// TIA Portal project "CHM_BORDEIRA_20190721" (V15)
// Frazer-Nash Consultancy Edits

(* hardware
DEVICE "SCALANCE X005"  SCALANCE X-Station
   slot 0: "SCALANCE X rack"  Rail
   slot 0: "Switch_1"  6GK5 008-0BA00-1AB2  V1.0
DEVICE "RIO 2/RIOCP-2T-ET 200iSP"  ET 200iSP station
   slot 0: "RIO 2 / RIOCP-2T"  Rail
   slot 2: "RIO 2 / RIOCP-2T - 5KF1 - IF Module"  ET200iSP  6ES7 152-1AA00-0AB0  V2.0
   slot 4: "6KF1 - 8DI x NAMUR"  8DI x NAMUR  6ES7 131-7RF00-0AB0
   slot 5: "7KF1 - 8DI x NAMUR"  8DI x NAMUR  6ES7 131-7RF00-0AB0
   slot 6: "8KF1 - 8DI x NAMUR"  8DI x NAMUR  6ES7 131-7RF00-0AB0
   slot 7: "9KF1 - 4DO x 23.1VDC / 20mA SD 'H'"  4DO x 23.1VDC / 20mA SD 'H'  6ES7 132-7RD01-0AB0
   slot 8: "10KF1 - 4AI x 2WIRE HART"  4AI x 2WIRE HART  6ES7 134-7TD00-0AB0
   slot 9: "11KF1 - 4AI x 2WIRE HART"  4AI x 2WIRE HART  6ES7 134-7TD00-0AB0
   slot 10: "12KF1 - 4AI x 2WIRE HART"  4AI x 2WIRE HART  6ES7 134-7TD00-0AB0
   slot 11: "13KF1 - 4AI x 2WIRE HART"  4AI x 2WIRE HART  6ES7 134-7TD00-0AB0
DEVICE "ET 200SP station_1"  ET 200SP-Station
   slot 0: "Rack_1"  Rack  6ES5 710-8MAx1
   slot 1: "Rack 1 - IGG PLC - 15KF2"  CPU 1510SP-1 PN  6ES7 510-1DJ01-0AB0  V2.1
   slot 2: "16KF1 - DI 16x24VDC ST_1"  DI 16x24VDC ST  6ES7 131-6BH00-0BA0  V1.1
      slot 1: "16KF1 - DI 16x24VDC ST_1"  DI 16x24VDC ST
   slot 3: "18KF1 - DI 16x24VDC ST_2"  DI 16x24VDC ST  6ES7 131-6BH00-0BA0  V1.1
      slot 1: "18KF1 - DI 16x24VDC ST_2"  DI 16x24VDC ST
   slot 4: "23KF1 - DQ 16x24VDC/0.5A ST_1"  DQ 16x24VDC/0.5A ST  6ES7 132-6BH00-0BA0  V1.1
      slot 1: "23KF1 - DQ 16x24VDC/0.5A ST_1"  DQ 16x24VDC/0.5A ST
   slot 5: "29KF1 - AI 8xI 2-,4-wire BA_1"  AI 8xI 2-,4-wire BA  6ES7 134-6GF00-0AA1  V1.0
      slot 1: "29KF1 - AI 8xI 2-,4-wire BA_1"  AI 8xI 2-,4-wire BA
   slot 6: "31KF1 - AI 8xI 2-,4-wire BA_2"  AI 8xI 2-,4-wire BA  6ES7 134-6GF00-0AA1  V1.0
      slot 1: "31KF1 - AI 8xI 2-,4-wire BA_2"  AI 8xI 2-,4-wire BA
   slot 7: "35KF1 - AQ 4xU/I ST_1"  AQ 4xU/I ST  6ES7 135-6HD00-0BA1  V1.1
      slot 1: "35KF1 - AQ 4xU/I ST_1"  AQ 4xU/I ST
   slot 8: "Server module_1"  Server module  6ES7 193-6PA00-0AA0  V1.0
      slot 1: "Server module_1"  Server module
   slot 127: "PROFINET BusAdapter CU"  BA 2xRJ45  6ES7 193-6AR00-0AA0  V0.0
      slot 32769: "Port_1"  6ES7 193-6AR00-0AA0
      slot 32770: "Port_2"  6ES7 193-6AR00-0AA0
DEVICE "ET 200SP station_2"  ET 200SP-Station
   slot 0: "Rack_2"  Rack  6ES5 710-8MAx1
   slot 1: "Rack 2 - BC PLC - 15KF3"  CPU 1510SP-1 PN  6ES7 510-1DJ01-0AB0  V2.1
   slot 2: "19KF1 - DI 16x24VDC ST_1"  DI 16x24VDC ST  6ES7 131-6BH00-0BA0  V1.1
      slot 1: "19KF1 - DI 16x24VDC ST_1"  DI 16x24VDC ST
   slot 3: "21KF1 - DI 16x24VDC ST_2"  DI 16x24VDC ST  6ES7 131-6BH00-0BA0  V1.1
      slot 1: "21KF1 - DI 16x24VDC ST_2"  DI 16x24VDC ST
   slot 4: "25KF1 - DQ 16x24VDC/0.5A ST_1"  DQ 16x24VDC/0.5A ST  6ES7 132-6BH00-0BA0  V1.1
      slot 1: "25KF1 - DQ 16x24VDC/0.5A ST_1"  DQ 16x24VDC/0.5A ST
   slot 5: "33KF1 - AI 8xI 2-,4-wire BA_1"  AI 8xI 2-,4-wire BA  6ES7 134-6GF00-0AA1  V1.0
      slot 1: "33KF1 - AI 8xI 2-,4-wire BA_1"  AI 8xI 2-,4-wire BA
   slot 6: "37KF1 - AQ 4xU/I ST_1"  AQ 4xU/I ST  6ES7 135-6HD00-0BA1  V1.1
      slot 1: "37KF1 - AQ 4xU/I ST_1"  AQ 4xU/I ST
   slot 7: "Server module_1"  Server module  6ES7 193-6PA00-0AA0  V1.0
      slot 1: "Server module_1"  Server module
   slot 127: "PROFINET BusAdapter CU"  BA 2xRJ45  6ES7 193-6AR00-0AA0  V0.0
      slot 32769: "Port_1"  6ES7 193-6AR00-0AA0
      slot 32770: "Port_2"  6ES7 193-6AR00-0AA0
DEVICE "S71500/ET200MP station_1"  S7-1500 station
   slot 0: "Rail_0"  Rack  6ES7 590-1***0-0AA0
   slot 1: "Rack 3 - GCU & BWT PLC - 7KF2"  CPU 1516F-3 PN/DP  6ES7 516-3FN01-0AB0  V2.1
      slot 3: "CPU display_1"  6ES7591-1BA00-0AA0
   slot 2: "8KF1 - DI 32x24VDC HF_1"  DI 32x24VDC HF  6ES7 521-1BL00-0AB0  V2.1
   slot 3: "12KF1 - DQ 32x24VDC/0.5A HF_1"  DQ 32x24VDC/0.5A HF  6ES7 522-1BL01-0AB0  V1.0
   slot 4: "16KF1 - AI 8xU/I HF_2"  AI 8xU/I HF  6ES7 531-7NF00-0AB0  V1.0
   slot 5: "18KF1 - AI 8xU/I HF_1"  AI 8xU/I HF  6ES7 531-7NF00-0AB0  V1.0
   slot 6: "20KF1 - AQ 4xU/I HF_1"  AQ 4xU/I HF  6ES7 532-5ND00-0AB0  V1.0
DEVICE "RIO 1/RIOCP-3T-ET 200iSP"  ET 200iSP station
   slot 0: "RIO 1 / RIOCP-3T"  Rail
   slot 2: "RIO 1 / RIOCP-3T - 5KF1 - IF Module"  ET200iSP  6ES7 152-1AA00-0AB0  V2.0
   slot 4: "6KF1 - 8DI x NAMUR_1"  8DI x NAMUR  6ES7 131-7RF00-0AB0
   slot 5: "7KF1 - 8DI x NAMUR_2"  8DI x NAMUR  6ES7 131-7RF00-0AB0
   slot 6: "8KF1 - 8DI x NAMUR_3"  8DI x NAMUR  6ES7 131-7RF00-0AB0
   slot 7: "9KF1 - 8DI x NAMUR_4"  8DI x NAMUR  6ES7 131-7RF00-0AB0
   slot 8: "10KF1 - 4DO x 23.1VDC / 20mA SD 'H'_1"  4DO x 23.1VDC / 20mA SD 'H'  6ES7 132-7RD01-0AB0
   slot 9: "11KF1 - 4DO x 23.1VDC / 20mA SD 'H'_2"  4DO x 23.1VDC / 20mA SD 'H'  6ES7 132-7RD01-0AB0
   slot 10: "12KF1 - 4AI x 2WIRE HART_1"  4AI x 2WIRE HART  6ES7 134-7TD00-0AB0
   slot 11: "13KF1 - 4AI x 2WIRE HART_2"  4AI x 2WIRE HART  6ES7 134-7TD00-0AB0
   slot 12: "14KF1 - 4AI x 2WIRE HART_1"  4AI x 2WIRE HART  6ES7 134-7TD00-0AB0
   slot 13: "15KF1 - 4AI x 2WIRE HART_2"  4AI x 2WIRE HART  6ES7 134-7TD00-0AB0
   slot 14: "16KF1 - 4AI x 2WIRE HART_3"  4AI x 2WIRE HART  6ES7 134-7TD00-0AB0
   slot 15: "17KF1 - 4AI x 2WIRE HART_4"  4AI x 2WIRE HART  6ES7 134-7TD00-0AB0
   slot 16: "Standby modules_1"  Standby modules  6ES7 138-7AA00-0AA0
DEVICE "RIO 3/RIOCP-2T-ET 200iSP"  ET 200iSP station
   slot 0: "RIO 3 / RIOCP-2T"  Rail
   slot 2: "RIO 3 / RIOCP-2T - 5KF1 - IF Module"  ET200iSP  6ES7 152-1AA00-0AB0  V2.0
   slot 4: "6KF1 - 8DI x NAMUR"  8DI x NAMUR  6ES7 131-7RF00-0AB0
   slot 5: "7KF1 - 8DI x NAMUR"  8DI x NAMUR  6ES7 131-7RF00-0AB0
   slot 6: "8KF1 - 8DI x NAMUR"  8DI x NAMUR  6ES7 131-7RF00-0AB0
   slot 7: "9KF1 - 4DO x 23.1VDC / 20mA SD 'H'"  4DO x 23.1VDC / 20mA SD 'H'  6ES7 132-7RD01-0AB0
   slot 8: "10KF1 - 4AI x 2WIRE HART_1"  4AI x 2WIRE HART  6ES7 134-7TD00-0AB0
   slot 9: "11KF1 - 4AI x 2WIRE HART"  4AI x 2WIRE HART  6ES7 134-7TD00-0AB0
   slot 10: "12KF1 - 4AI x 2WIRE HART"  4AI x 2WIRE HART  6ES7 134-7TD00-0AB0
   slot 11: "13KF1 - 4AI x 2WIRE HART"  4AI x 2WIRE HART  6ES7 134-7TD00-0AB0
DEVICE "RIO 4/RIOCP-2T-ET 200iSP"  ET 200iSP station
   slot 0: "RIO 4 / RIOCP-2T"  Rail
   slot 2: "RIO 4 / RIOCP-2T - 5KF1 - IF Module"  ET200iSP  6ES7 152-1AA00-0AB0  V2.0
   slot 4: "6KF1 - 8DI x NAMUR"  8DI x NAMUR  6ES7 131-7RF00-0AB0
   slot 5: "7KF1 - 8DI x NAMUR"  8DI x NAMUR  6ES7 131-7RF00-0AB0
   slot 6: "8KF1 - 8DI x NAMUR"  8DI x NAMUR  6ES7 131-7RF00-0AB0
   slot 7: "9KF1 - 4DO x 23.1VDC / 20mA SD 'H'"  4DO x 23.1VDC / 20mA SD 'H'  6ES7 132-7RD01-0AB0
   slot 8: "10KF1 - 4AI x 2WIRE HART_1"  4AI x 2WIRE HART  6ES7 134-7TD00-0AB0
   slot 9: "11KF1 - 4AI x 2WIRE HART_1"  4AI x 2WIRE HART  6ES7 134-7TD00-0AB0
   slot 10: "12KF1 - 4AI x 2WIRE HART"  4AI x 2WIRE HART  6ES7 134-7TD00-0AB0
   slot 11: "13KF1 - 4AI x 2WIRE HART"  4AI x 2WIRE HART  6ES7 134-7TD00-0AB0
DEVICE "RIO 5/RIOCP-2T-ET 200iSP"  ET 200iSP station
   slot 0: "RIO 5 / RIOCP-2T"  Rail
   slot 2: "RIO 5 / RIOCP-2T - 5KF1 - IF Module"  ET200iSP  6ES7 152-1AA00-0AB0  V2.0
   slot 4: "6KF1 - 8DI x NAMUR_1"  8DI x NAMUR  6ES7 131-7RF00-0AB0
   slot 5: "7KF1 - 8DI x NAMUR_2"  8DI x NAMUR  6ES7 131-7RF00-0AB0
   slot 6: "8KF1 - 8DI x NAMUR_3"  8DI x NAMUR  6ES7 131-7RF00-0AB0
   slot 7: "9KF1 - 4DO x 23.1VDC / 20mA SD 'H'_1"  4DO x 23.1VDC / 20mA SD 'H'  6ES7 132-7RD01-0AB0
   slot 8: "10KF1 - 4AI x 2WIRE HART_1"  4AI x 2WIRE HART  6ES7 134-7TD00-0AB0
   slot 9: "11KF1- 4AI x 2WIRE HART_1"  4AI x 2WIRE HART  6ES7 134-7TD00-0AB0
   slot 10: "12KF1 - 4AI x 2WIRE HART_2"  4AI x 2WIRE HART  6ES7 134-7TD00-0AB0
   slot 11: "13KF1 - 4AI x 2WIRE HART_3"  4AI x 2WIRE HART  6ES7 134-7TD00-0AB0
DEVICE "RIO 7/RIOCP-1T-ET 200iSP"  ET 200iSP station
   slot 0: "RIO 7/ RIOCP-1T"  Rail
   slot 2: "RIO 7 / RIOCP-1T - 5KF1 - IF Module"  ET200iSP  6ES7 152-1AA00-0AB0  V2.0
   slot 4: "6KF1 - 8DI x NAMUR"  8DI x NAMUR  6ES7 131-7RF00-0AB0
   slot 5: "7KF1 - 8DI x NAMUR"  8DI x NAMUR  6ES7 131-7RF00-0AB0
   slot 6: "8KF1 - 4DO x 23.1VDC / 20mA SD 'H'_1"  4DO x 23.1VDC / 20mA SD 'H'  6ES7 132-7RD01-0AB0
   slot 7: "9KF1 - 4AI x 2WIRE HART_1"  4AI x 2WIRE HART  6ES7 134-7TD00-0AB0
   slot 8: "10KF1 - 4AI x 2WIRE HART"  4AI x 2WIRE HART  6ES7 134-7TD00-0AB0
   slot 9: "11KF1 - 4AI x 2WIRE HART"  4AI x 2WIRE HART  6ES7 134-7TD00-0AB0
DEVICE "RIO 6/RIOCP-2T-ET 200iSP"  ET 200iSP station
   slot 0: "RIO 6 / RIOCP-2T"  Rail
   slot 2: "RIO 6 / RIOCP-2T - 5KF1 - IF Module"  ET200iSP  6ES7 152-1AA00-0AB0  V2.0
   slot 4: "6KF1 - 8DI x NAMUR_1"  8DI x NAMUR  6ES7 131-7RF00-0AB0
   slot 5: "7KF1 - 8DI x NAMUR_2"  8DI x NAMUR  6ES7 131-7RF00-0AB0
   slot 6: "8KF1 - 8DI x NAMUR_3"  8DI x NAMUR  6ES7 131-7RF00-0AB0
   slot 7: "9KF1 - 4DO x 23.1VDC / 20mA SD 'H'_1"  4DO x 23.1VDC / 20mA SD 'H'  6ES7 132-7RD01-0AB0
   slot 8: "10KF1 - 4AI x 2WIRE HART_1"  4AI x 2WIRE HART  6ES7 134-7TD00-0AB0
   slot 9: "11KF1- 4AI x 2WIRE HART_1"  4AI x 2WIRE HART  6ES7 134-7TD00-0AB0
   slot 10: "12KF1 - 4AI x 2WIRE HART_2"  4AI x 2WIRE HART  6ES7 134-7TD00-0AB0
   slot 11: "13KF1 - 4AI x 2WIRE HART_3"  4AI x 2WIRE HART  6ES7 134-7TD00-0AB0
DEVICE "IGG HMI"  TP1500 Comfort
   slot 0: "IGG HMI"  TP1500 Comfort  6AV2 124-0QC02-0AX0  15.0.0.0
   slot 1: "HMI_RT_1"  TP1500 Comfort  6AV2 124-0QC02-0AX0  15.0.0.0
   slot 5: "IGG HMI.IE_CP_1"  PROFINET Interface  15.0.0.0
      slot 1: "PROFINET Interface_1"  PROFINET Interface
         slot 1: "Port_1"  Port
         slot 2: "Port_2"  Port
   slot 6: "IGG HMI.IE_CP_2"  PROFINET Interface  15.0.0.0
      slot 1: "PROFINET Interface_GBit"  PROFINET Interface
         slot 1: "Port_1"  Port
   slot 7: "IGG HMI.MPI/DP_CP_1"  MPI/DP Interface  15.0.0.0
DEVICE "CCR HMI"  TP1200 Comfort
   slot 0: "CCR HMI"  TP1200 Comfort  6AV2 124-0MC01-0AX0  15.0.0.0
   slot 1: "HMI_RT_4"  TP1200 Comfort  6AV2 124-0MC01-0AX0  15.0.0.0
   slot 5: "CCR HMI._CP_1"  PROFINET Interface  15.0.0.0
      slot 1: "PROFINET Interface_1"  PROFINET Interface
         slot 1: "Port_1"  Port
         slot 2: "Port_2"  Port
   slot 7: "CCR HMI.I/DP_CP_1"  MPI/DP Interface  15.0.0.0
DEVICE "Bridge HMI"  KTP400 Comfort
   slot 0: "Bridge HMI"  KTP400 Comfort  6AV2 124-2DC01-0AX0  15.0.0.0
   slot 1: "HMI_RT_2"  KTP400 Comfort  6AV2 124-2DC01-0AX0  15.0.0.0
   slot 5: "Bridge HMI.1"  PROFINET Interface  15.0.0.0
      slot 1: "PROFINET Interface_1"  PROFINET Interface
         slot 1: "Port_1"  Port
   slot 7: "Bridge HMI._CP_1"  MPI/DP Interface  15.0.0.0
DEVICE "GSD device_1"  GSD.Device.PN
   slot 0: "Rack"  Rack  V1.0
   slot 0: "WBT"  Serial  HD674-A006
      slot 0: "Submodule V1"  Submodule V1
      slot 1: "I"  I
         slot 1: "P1"  P1
         slot 2: "P2"  P2
   slot 1: "IO"  Module  12345-0040-M
      slot 0: "Module"  Module
*)

// ===== PLC "Rack 1 - IGG PLC - 15KF2"  CPU 1510SP-1 PN =====

VAR_GLOBAL   // PLC tag table "Default tag table"
   "System_Byte" AT %MB1 : Byte;
   "FirstScan" AT %M1.0 : Bool;
   "DiagStatusUpdate" AT %M1.1 : Bool;
   "AlwaysTRUE" AT %M1.2 : Bool;
   "AlwaysFALSE" AT %M1.3 : Bool;
   "Clock_Byte" AT %MB0 : Byte;
   "Clock_10Hz" AT %M0.0 : Bool;
   "Clock_5Hz" AT %M0.1 : Bool;
   "Clock_2.5Hz" AT %M0.2 : Bool;
   "Clock_2Hz" AT %M0.3 : Bool;
   "Clock_1.25Hz" AT %M0.4 : Bool;
   "Clock_1Hz" AT %M0.5 : Bool;
   "Clock_0.625Hz" AT %M0.6 : Bool;
   "Clock_0.5Hz" AT %M0.7 : Bool;
   "IGG E-Stop Healthy" AT %I0.0 : Bool;   // S2-8K1
   "CA Blower Ready" AT %I0.1 : Bool;   // E139-MCCP/6TA1
   "Fuel Pump 1 Tripped" AT %I0.2 : Bool;   // E500A-MCCP/7Q2
   "Fuel Pump 2 Tripped" AT %I0.3 : Bool;   // E500B-MCCP/7Q3
   "Fuel Pump 1 Enabled" AT %I0.4 : Bool;   // E500A-MCCP/9Q1
   "Fuel Pump 2 Enabled" AT %I0.5 : Bool;   // E500B-MCCP/9Q2
   "IG Supply Valve Opened" AT %I0.6 : Bool;   // CV401-16B1
   "IG Supply Valve Closed" AT %I0.7 : Bool;   // CV401-16B1
   "DTB Valve Opened" AT %I1.0 : Bool;   // CV321-17B1
   "DTB Valve Closed" AT %I1.1 : Bool;   // CV321-17B1
   "CSW Drain Valve Opened" AT %I1.2 : Bool;   // CV322-17B2
   "CSW Drain Valve Closed" AT %I1.3 : Bool;   // CV322-17B2
   "CSW Valve Open" AT %I1.4 : Bool;   // CV311-17B3
   "CSW Valve Closed" AT %I1.5 : Bool;   // CV311-17B3
   "Flue Gas Scrubber CSW Valve Opened" AT %I1.6 : Bool;   // CV312-17B4
   "Flue Gas Scrubber CSW Valve Closed" AT %I1.7 : Bool;   // CV312-17B4
   "BC PLC Power Healthy" AT %I2.0 : Bool;   // -15Q4
   "IGG Vent Power Healthy" AT %I2.1 : Bool;   // -6Q2
   "MCC Vent Power Healthy" AT %I2.2 : Bool;   // -MCCP/8Q4
   "7T1 Power Healthy" AT %I2.3 : Bool;   // -7T1 Controls Power
   "7T2 Power Healthy" AT %I2.4 : Bool;   // -7T2 IGG Power
   "7T3 Power Healthy" AT %I2.5 : Bool;   // -7T3 BC Power
   "Maintained 24V Power" AT %I2.6 : Bool;   // -7Q4
   "Safety System Interlock" AT %I2.7 : Bool;   // Safety interlock
   "Cargo Blanketing IG Supply Valve Open" AT %I3.0 : Bool;   // CV431-25QM8
   "Cargo Blanketing IG Supply Valve Close" AT %I3.1 : Bool;   // CV431-25QM8
   "BWTS IG Supply Valve Open" AT %I3.2 : Bool;   // CV432-25QM8
   "BWTS IG Supply Valve Close" AT %I3.3 : Bool;   // CV432-25QM8
   "CA Blower Running" AT %I3.4 : Bool;   // E139-MCCP/6TA1
   "VSD Fault" AT %I3.5 : Bool;   // E139-MCCP/6TA1
   "Correct Phase Rotation" AT %I3.6 : Bool;   // -MCCP/5PG1
   "R1_SPR_DI_3_7" AT %I3.7 : Bool;   // Spare input
   "CA Pressure PIT102" AT %IW112 : Int;   // PIT102-29B1
   "IG Temp" AT %IW114 : Int;   // TIT401-29B2
   "IG Outlet Pressure PIT402" AT %IW116 : Int;   // PIT402-29B3
   "IG Vent Valve Position Feedback" AT %IW118 : Int;   // CV403-29B4
   "CA Blower RPM" AT %IW120 : Int;   // E139-6TA1
   "CA Blower Current" AT %IW122 : Int;   // E139-6TA1
   "FW Bulk Tank Level Transmitter" AT %IW124 : Int;   // LIT305
   "Atm Oxygen Content 1" AT %IW128 : Int;   // Crowcon Atmospheric Sensors-31B1
   "Atm Oxygen Content 2" AT %IW130 : Int;   // Crowcon Atmospheric Sensors-31B2
   "R1_SPR_AI_132" AT %IW132 : Int;   // Spare
   "Shell CSW Temp TIT315" AT %IW134 : Int;   // TIT315-31B4
   "Inlet CSW Temp TIT319" AT %IW136 : Int;   // TIT319-32B1
   "Outlet CSW Temp TIT360" AT %IW138 : Int;   // TIT360-32B2
   "Inlet CSW Pressure PIT359" AT %IW140 : Int;   // PIT359-32B3
   "Outlet CSW Pressure PIT316" AT %IW142 : Int;   // PIT316-32B4
   "Fuel Pump 1 Control" AT %Q0.0 : Bool;   // E500-MCCP/9Q1
   "Fuel Pump 2 Control" AT %Q0.1 : Bool;   // E500-MCCP/9Q1
   "CA Blower Control" AT %Q0.2 : Bool;   // E139-MCCP/6TA1
   "CSW Inlet Valves Control" AT %Q0.3 : Bool;   // CV311/CV312-23QM1
   "CSW Drain Valves Control" AT %Q0.4 : Bool;   // CV321/CV322-23QM2
   "IG Supply Valve Control" AT %Q0.5 : Bool;   // CV401
   "R1_SPR_DQ_1_0" AT %Q1.0 : Bool;   // Spare input
   "Atmospheric Alarm" AT %Q1.1 : Bool;   // -24K2
   "IGG Shutdown Alarm Active" AT %Q1.2 : Bool;   // -24K3
   "IGG Warning Alarm Active" AT %Q1.3 : Bool;   // -24K4
   "IGG Running" AT %Q1.4 : Bool;   // -24PF1
   "Shutdown Alarm" AT %Q1.5 : Bool;   // -24PF2
   "Warning Alarm" AT %Q1.6 : Bool;   // -24PF3
   "Buzzer" AT %Q1.7 : Bool;   // -24PF4
   "Vent Valve Position Control" AT %QW98 : Int;   // CV403-35QN1
   "R1_SPR_AI_126" AT %IW126 : Int;   // Spare input
   "Cargo Blanketing/BWTS Valve Control" AT %Q0.6 : Bool;   // CV431/432-25QM8
   "R1_SPR_DQ_0_7" AT %Q0.7 : Bool;   // Spare input
   "CA Blower Speed Control" AT %QW100 : Word;   // E139-MCCP/6TA1
   "R1_SPR_AQ_102" AT %QW102 : Word;   // Spare output
   "R1_SPR_AQ_104" AT %QW104 : Word;   // Spare output
   "db_time_sync_time_system_READ" AT %M2.0 : LDT;
   "db_time_sync_time_local_READ" AT %M4.0 : LDT;
   "TimeRetVal1" AT %MW8 : Int;
   "RESET_STEP" AT %M12.0 : Bool;
   "IGG_ALARM_ACKNLG_1" AT %MW12 : Word;   // %MW12.DBX0.0
   "IGG_ALARM_ACKNLG_2" AT %MW14 : Word;
   "IGG_ALARM_ACKNLG_3" AT %MW16 : Word;
   "IGG_ALARM_ACKNLG_4" AT %MW18 : Word;
   "IGG_ALARM_ACKNLG_5" AT %MW20 : Word;
   "IGG_ALARM_ACKNLG_6" AT %MW22 : Word;
   "BC_ALARM_ACKNLG_1" AT %MW24 : Word;
   "BC_ALARM_ACKNLG_2" AT %MW26 : Word;
   "BC_ALARM_ACKNLG_3" AT %MW28 : Word;
   "BC_ALARM_ACKNLG_4" AT %MW30 : Word;
   "BC_ALARM_ACKNLG_5" AT %MW32 : Word;
   "BC_ALARM_ACKNLG_6" AT %MW34 : Word;
   "Tag_1" AT %M233.3 : Bool;
   "Tag_2" AT %M233.4 : Bool;
   "Tag_3" AT %M233.5 : Bool;
   "Tag_4" AT %M233.6 : Bool;
   "Tag_5" AT %M233.7 : Bool;
END_VAR

TYPE "AI_Data"
VERSION : 0.1
   STRUCT
      RAW_MIN : Int;   // Raw minimum value from AI card
      RAW_MAX : Int := 27648;   // Raw maximum value from AI card
      NORM : Real;   // Normalised real value
      ENG_MIN : Real;   // Engineering units minimum value
      ENG_MAX : Real := 100.0;   // Engineering units maximum value
   END_STRUCT;
END_TYPE

TYPE "AQ_Data"
VERSION : 0.1
   STRUCT
      ENG_MIN : Real;   // Engineering units minimum value
      ENG_MAX : Real := 100.0;   // Engineering units maximum value
      NORM : Real;   // Normalised real value
      RAW_MIN : Int;   // Raw minimum value from AQ card
      RAW_MAX : Int := 27648;   // Raw maximum value from AQ card
   END_STRUCT;
END_TYPE

// folder: 10 - 19 IO & Processing

DATA_BLOCK "Alarm beacon handling_DB"   // DB1
{ S7_Optimized_Access := 'TRUE' }
VERSION : 0.1
// stored: InstanceOfName Alarm beacon handling
"Alarm beacon handling"
BEGIN
END_DATA_BLOCK

DATA_BLOCK "Date_And_Time_Data"   // DB3
{ S7_Optimized_Access := 'TRUE' }
VERSION : 0.1
   VAR
      SYSTEM_TIME : DTL;
      LOCAL_TIME : DTL;
      HMI_INPUT_FIELD_TIME_IGG : DTL;
      SYNCH_HMI_CLOCK_IGG : Bool;
      GET_TIME_IGG : Bool;
      HMI_INPUT_FIELD_TIME_CCR : DTL;
      SYNCH_HMI_CLOCK_CCR : Bool;
      GET_TIME_CCR : Bool;
   END_VAR
BEGIN
END_DATA_BLOCK

DATA_BLOCK "10_DI_Data"   // DB10
TITLE = Digital Input Data
{ S7_Optimized_Access := 'TRUE' }
AUTHOR : JRS
VERSION : 0.1
// Processed data for code use
   VAR
      IGG_ESTOP_OK : Bool;   // IGG E-Stop healthy (S2-8K1)
      BC_PLC_PWR_OK : Bool;   // BC PLC Power healthy
      IGG_VNT_PWR_OK : Bool;   // IGG Vent power healthy
      MCC_VNT_PWR_OK : Bool;   // MCC Vent power healthy
      "7T1_PWR_OK" : Bool;   // 7T1 Power healthy
      "7T2_PWR_OK" : Bool;   // 7T2 Power healthy
      "7T3_PWR_OK" : Bool;   // 7T3 Power healthy
      MAINTD_24VDC_PWR_OK : Bool;   // Maintained 24V power
      SFTY_SYS_IL : Bool;   // Safety system interlock
      R1_SPR_DI_3_7 : Bool;   // Spare input
      MCCP_5PG1_OK : Bool;   // Correct phase rotation
      CV311_OPN : Bool;   // CSW Valve Open
      CV311_CLSD : Bool;   // CSW Valve Closed
      CV312_OPN : Bool;   // Flue Gas Scrubber CSW valve open
      CV312_CLSD : Bool;   // Flue gas scrubber CSW valve closed
      CV321_OPN : Bool;   // DTB valve open
      CV321_CLSD : Bool;   // DTB valve closed
      CV322_OPN : Bool;   // CSW Drain valve open
      CV322_CLSD : Bool;   // CSW drain valve closed
      CV401_OPN : Bool;   // IG supply valve open
      CV401_CLSD : Bool;   // IG supply valve closed
      CV431_OPN : Bool;   // Cargo blanketing IG supply valve open
      CV431_CLSD : Bool;   // Cargo blanketing IG supply valve closed
      CV432_OPN : Bool;   // BWTS IG supply valve open
      CV432_CLSD : Bool;   // BWTS IG supply valve closed
      E139_READY : Bool;   // CA blower ready
      E139_RUNNING : Bool;   // CA blower running
      E139_VSD_FLT : Bool;   // CA blower VSD fault
      E500A_ENBLD : Bool;   // Fuel pump 1 enabled
      E500A_TRIPPED : Bool;   // Fuel pump 1 tripped
      E500B_ENBLD : Bool;   // Fuel pump 2 enabled
      E500B_TRIPPED : Bool;   // Fuel pump 2 tripped
   END_VAR
BEGIN
END_DATA_BLOCK

DATA_BLOCK "12_AI_Data"   // DB12
TITLE = Analogue Input Data
{ S7_Optimized_Access := 'TRUE' }
AUTHOR : JRS
VERSION : 0.1
// Processed data for code use
   VAR
      PIT102_SCALED : Real;   // CA Pressure
      TIT401_SCALED : Real;   // IG Temperature
      PIT402_SCALED : Real;   // IG Outlet pressure
      CV403_SCALED : Real;   // IG Vent position feedback
      E139_RPM_SCALED : Real;   // CA Blower RPM
      E139_AMPS_SCALED : Real;   // CA Blower current
      LIT305_SCALED : Real;   // FW Bulk tank level
      R1_SPR_AI_126_SCALED : Real;   // Spare input
      R1_SPR_AI_132_SCALED : Real;   // Spare input
      AT_O2_01_SCALED : Real;   // Atmospheric oxygen content 1
      AT_O2_02_SCALED : Real;   // Atmospheric oxygen content 2
      TIT315_SCALED : Real;   // CSW Temperature at IGG shell
      TIT319_SCALED : Real;   // CSW Temperature at IGG inlet
      TIT360_SCALED : Real;   // CSW Temperature at IGG outlet
      PIT359_SCALED : Real;   // CSW Pressure at IGG inlet
      PIT316_SCALED : Real;   // CSW Pressure at IGG outlet
      IW_112 : "AI_Data";   // PIT102 calibration data
      IW_114 : "AI_Data";   // TIT401 calibration data
      IW_116 : "AI_Data";   // PIT402 calibration data
      IW_118 : "AI_Data";   // CV403 calibration data
      IW_120 : "AI_Data";   // E139 Running Speed calibration data
      IW_122 : "AI_Data";   // E139 Current calibration data
      IW_124 : "AI_Data";   // LIT305 calibration data
      IW_126 : "AI_Data";   // Spare input calibration data
      IW_128 : "AI_Data";   // 31B1 calibration data
      IW_130 : "AI_Data";   // 31B2 calibration data
      IW_132 : "AI_Data";   // Spare input calibration data
      IW_134 : "AI_Data";   // TIT315 calibration data
      IW_136 : "AI_Data";   // TIT319 calibration data
      IW_138 : "AI_Data";   // TIT360 calibration data
      IW_140 : "AI_Data";   // PIT359 calibration data
      IW_142 : "AI_Data";   // PIT316 calibration data
   END_VAR
BEGIN
   IW_114.ENG_MAX := 150.0;   // Engineering units maximum value - degC
   IW_112.ENG_MAX := 1000.0;   // Engineering units maximum value - bar(g)
   IW_116.ENG_MAX := 1000.0;   // Engineering units maximum value - bar(g)
   IW_136.ENG_MIN := 0.0;   // Engineering units minimum value - degC
   IW_134.ENG_MIN := 0.0;   // Engineering units minimum value - degC
   IW_128.ENG_MAX := 25.0;
   IW_130.ENG_MAX := 25.0;
   IW_132.ENG_MAX := 40.0;
   IW_134.ENG_MAX := 150.0;   // Engineering units maximum value - degC
   IW_136.ENG_MAX := 150.0;   // Engineering units maximum value - degC
   IW_138.ENG_MAX := 150.0;   // Engineering units maximum value - degC
   IW_140.ENG_MAX := 10.0;   // Engineering units maximum value - bar(g)
   IW_142.ENG_MAX := 10.0;   // Engineering units maximum value - bar(g)
   IW_112.ENG_MIN := 0.0;   // Engineering units minimum value - bar(g)
   IW_114.ENG_MIN := 0.0;   // Engineering units minimum value - degC
   IW_116.ENG_MIN := 0.0;   // Engineering units minimum value - bar(g)
   IW_118.ENG_MIN := 0.0;   // Engineering units minimum value (%)
   IW_118.ENG_MAX := 100.0;   // Engineering units maximum value (%)
   IW_138.ENG_MIN := 0.0;   // Engineering units minimum value - degC
   IW_140.ENG_MIN := 0.0;   // Engineering units minimum value - bar(g)
   IW_142.ENG_MIN := 0.0;   // Engineering units minimum value - bar(g)
   IW_122.ENG_MAX := 100.0;
   IW_120.ENG_MAX := 1782.0;
END_DATA_BLOCK

DATA_BLOCK "14_DQ_Data"   // DB14
TITLE = Digital Output Data
{ S7_Optimized_Access := 'TRUE' }
AUTHOR : JRS
VERSION : 0.1
// Processed data for output via physical connection
   VAR
      E500A_CNTRL : Bool;   // Run fuel pump #1
      E500B_CNTRL : Bool;   // Run fuel pump #2
      CV311_312_CNTRL : Bool;   // CSW Inlet valves control
      CV321_322_CNTRL : Bool;   // CSW Outlet valves control
      CV401_CNTRL : Bool;   // IG Supply valve control
      E139_CNTRL : Bool;   // Run combustion air blower
      CV431_432_CNTRL : Bool;   // Cargo blanketting/BWTS valve control
      "24K2" : Bool;   // Atmospheric alarm
      "24K3" : Bool;   // IGG Shutdown alarm active
      "24K4" : Bool;   // IGG Warning alarm active
      "24PF1" : Bool;   // IGG Running
      "24PF2" : Bool;   // Shutdown alarm
      "24PF3" : Bool;   // Warning alarm
      "24PF4" : Bool;   // Buzzer
      R2_SPR_DQ_0_7 : Bool;   // Spare output
      R2_SPR_DQ_1_0 : Bool;   // Spare output
   END_VAR
BEGIN
END_DATA_BLOCK

DATA_BLOCK "16_AQ_Data"   // DB16
TITLE = Analogue Output Data
{ S7_Optimized_Access := 'TRUE' }
AUTHOR : JRS
VERSION : 0.1
// Processed data for output via physical connection
   VAR RETAIN
      CV403_CNTRL : Real;   // Vent position control
      E139_SPEED : Real;   // CA Blower speed control
   END_VAR
   VAR
      R1_SPR_AQ_102 : Real;   // Spare output
      R1_SPR_AQ_104 : Real;   // Spare output
      QW_98 : "AQ_Data";   // CV403 calibration data
      QW_100 : "AQ_Data";   // E139 Speed Control calibration data
      QW_102 : "AQ_Data";   // Spare output calibration data
      QW_104 : "AQ_Data";   // Spare output calibration data
   END_VAR
BEGIN
   QW_98.ENG_MIN := 0.0;   // Engineering units minimum value - %
   QW_98.ENG_MAX := 100.0;   // Engineering units maximum value - %
   QW_100.ENG_MIN := 0.0;
   QW_100.ENG_MAX := 1782.0;
END_DATA_BLOCK

DATA_BLOCK "19_AUTO_CMNDS_Data"   // DB19
TITLE = Automatic Commands Data
{ S7_Optimized_Access := 'TRUE' }
AUTHOR : JRS
VERSION : 0.1
// Defined data for use prior to output processing
   VAR
      Fuel_Pump_Demand : Bool;   // 1 = Run, 0 = Not
      PIT402_Ramp_Demand : Bool;   // 1 = Run, 0 = Not
      CV403_PID_MDLTG : Bool;   // 1 = Modulating, 0 = Not
      ALRM_EDGE : Bool;   // Pulse bit
      PIT402_Target : Real := 40.0;   // PIT402 burner target setpoint (bar g)
      PIT402_LowLow : Real := 30.0;   // PIT402 burner low low setpoint (bar g)
      PIT402_Low : Real := 35.0;   // PIT402 burner low setpoint (bar g)
      PIT402_High : Real := 80.0;   // PIT402 burner high setpoint (bar g)
      PIT402_HighHigh : Real := 100.0;   // PIT402 burner high high setpoint (bar g)
      PIT102_LowLow : Real := 30.0;   // PIT102 burner low low setpoint (bar g)
      PIT102_Low : Real := 35.0;   // PIT102 burner low setpoint (bar g)
      PIT102_High : Real := 80.0;   // PIT102 burner high setpoint (bar g)
      PIT102_HighHigh : Real := 100.0;   // PIT102 burner high high setpoint (bar g)
   END_VAR
BEGIN
END_DATA_BLOCK

DATA_BLOCK "Evolving Setpoint_DB20"   // DB20
{ S7_Optimized_Access := 'TRUE' }
VERSION : 0.1
// stored: InstanceOfName Evolving Setpoint
"Evolving Setpoint"
BEGIN
END_DATA_BLOCK

// folder: 100 - 119 Automatic Functions

DATA_BLOCK "100_IGG_AUTO_SEQ_DB"   // DB100
TITLE = IGG Auto Sequence Instance DB
{ S7_Optimized_Access := 'TRUE' }
AUTHOR : JRS
VERSION : 0.1
// Data required for FB
// stored: InstanceOfName 100_IGG_AUTO_SEQ
"100_IGG_AUTO_SEQ"
BEGIN
END_DATA_BLOCK

DATA_BLOCK "101_Fuel_Pumps_DB"   // DB101
TITLE = Fuel Pumps Instance DB
{ S7_Optimized_Access := 'TRUE' }
AUTHOR : JRS
VERSION : 0.1
// Data required for FB
// stored: InstanceOfName 101_Fuel_Pumps
"101_Fuel_Pumps"
BEGIN
END_DATA_BLOCK

DATA_BLOCK "105_SP_RAMP_PIT402_UP_DB"   // DB105
{ S7_Optimized_Access := 'TRUE' }
AUTHOR : JRS
VERSION : 0.1
// stored: InstanceOfName 105_SP_RAMP_PIT402_UP
"105_SP_RAMP_PIT402_UP"
BEGIN
END_DATA_BLOCK

DATA_BLOCK "107_SP_RAMP_PIT402_DN_DB"   // DB107
{ S7_Optimized_Access := 'TRUE' }
AUTHOR : JRS
VERSION : 0.1
// stored: InstanceOfName 107_SP_RAMP_PIT402_DN
"107_SP_RAMP_PIT402_DN"
BEGIN
END_DATA_BLOCK

// folder: 120 - 139 FAT Functions

DATA_BLOCK "120_FAT_FCS_DB"   // DB120
TITLE = FAT Functions Data Area
{ S7_Optimized_Access := 'TRUE' }
AUTHOR : JRS
VERSION : 0.1
// For data relating to the FAT mode and functionality
   VAR
      IN_FAT : Bool;   // In FAT mode
      INTO_FAT_PLS : Bool;   // Pulse bit
      INTO_FAT_TMD_PLS : TP_TIME;   // Into FAT pulse timer
   END_VAR
BEGIN
   INTO_FAT_TMD_PLS.PT := T#100ms;
END_DATA_BLOCK

// folder: 300 - 499 Counters and Timer DBs

DATA_BLOCK "300_AUT_SEQ_TMRS_DB"   // DB300
TITLE = Auto Sequence Timers Data
{ S7_Optimized_Access := 'TRUE' }
AUTHOR : JRS
VERSION : 0.1
// Data area for auto sequence timers
   VAR RETAIN
      PRE_BC_STRT_CMND_DLY : TON_TIME;   // For the delay prior to the BC start command
      PRE_CV203_CLS_CMND_DLY : TON_TIME;   // For the delay prior to the CV203 close command
      POST_P301_STOP_DLY : TON_TIME;   // For the delay after P301 stopped
      POST_CV311_CLS_DLY : TON_TIME;   // For the delay after CV311 closed
      POST_CV311_CLS_DLY_1 : TON_TIME;
      POST_CV321_OPN_DLY : TON_TIME;   // For the delay after CV321 opened
      "NOK INTLK DLY" : TON_TIME;   // Interlocks not OK delay
      "E500 A Ctrl Delay" : TON_TIME;
      "E500 B Ctrl Delay" : TON_TIME;
      "E500 A Enable Delay" : TOF_TIME;
      "E500 B Enable Delay" : TOF_TIME;
      "CV127_CLOSED Delay" : TON_TIME;
      "E139 Start Check Delay" : TON_TIME;
   END_VAR
   VAR
      "E139 RUNNING Delay" : TON_TIME;
   END_VAR
   VAR RETAIN
      "P301 CSW Pump Delay after start" : TON_TIME;
      "ALARM STOP" : TP_TIME;
      "Pilot Burner Purge Stage Complete" : TON_TIME;
   END_VAR
   VAR
      "Pilot Burner Purge Stage Complete_TOF" : TOF_TIME;
      "Cooling System Overrun CV311" : TOF_TIME;
      "Cooling System Overrun CV321" : TOF_TIME;
      "Cooling System Overrun P301" : TOF_TIME;
      "STEP190 Delay Post Burn" : TON_TIME;
      "E500A Trip Delay" : TON_TIME;
      "E500B Trip Delay" : TON_TIME;
      "STOP Puls" : TP_TIME;
      "E-Stop BWT" : TOF_TIME;
      "E-Stop Delay for CSW Inlet" : TOF_TIME;
      "E-Stop Delay for CSW Outlet" : TOF_TIME;
      "CSW OVR Outlet Stop Delay" : TON_TIME;
   END_VAR
BEGIN
   PRE_BC_STRT_CMND_DLY.PT := T#10s;
   "NOK INTLK DLY".PT := T#3s;
   "E500 A Ctrl Delay".PT := T#2s;
   "E500 B Ctrl Delay".PT := T#2s;
   "E139 Start Check Delay".PT := T#15s;
   "P301 CSW Pump Delay after start".PT := T#5s;
   PRE_CV203_CLS_CMND_DLY.PT := T#3s;
   POST_P301_STOP_DLY.PT := T#3s;
   POST_CV311_CLS_DLY.PT := T#3s;
   POST_CV311_CLS_DLY_1.PT := T#3s;
   POST_CV321_OPN_DLY.PT := T#3s;
   "E500 A Enable Delay".PT := T#1s;
   "E500 B Enable Delay".PT := T#1s;
   "CV127_CLOSED Delay".PT := T#3s;
   "E500A Trip Delay".PT := T#1s;
   "E500B Trip Delay".PT := T#1s;
   "E-Stop BWT".PT := T#1s;
   "E-Stop Delay for CSW Inlet".PT := T#30s;
   "E-Stop Delay for CSW Outlet".PT := T#40s;
   "CSW OVR Outlet Stop Delay".PT := T#30s;
END_DATA_BLOCK

// folder: 50 - 59 Communication

DATA_BLOCK "50_CMND_DATA"   // DB50
TITLE = Command Data
{ S7_Optimized_Access := 'FALSE' }
AUTHOR : JRS
VERSION : 0.1
// Data area for commands from master PLC
   VAR
      HEART_BEAT : Bool;   // Heartbeat
      CRNT_MODE : Int := 1;   // 1 = Auto, 2 = Man, 3 = FatAuto, 4 = FatMan
      RST_AUT_SEQ : Bool;   // Reset automatic sequence
      GCU_BWT_ALARM : Bool;   // 1 = Alarm, 0 = Not
      OK_RUN_IGG : Bool;   // 1 = Run IGG, 0 = Not
      STOP_IGG : Bool;   // 1 = Stop IGG, 0 = Not
      OPEN_CV401 : Bool;   // 1 = Open, 0 = Not
      RUN_P305 : Bool;   // 1 = Run pump, 0 = Not
      GCU_WRNG_ACTV : Bool;   // 1 = GCU Warning active, 0 = Not
      SPR_BOOL : Bool;   // Spare bit
      RUN_P301 : Bool;   // 1 = Run pump, 0 = Not
      OPEN_CV311 : Bool;   // 1 = Open, 0 = Not
      OPEN_CV322 : Bool;   // 1 = Open, 0 = Not
      NewALARM : Bool;   // NewALARM
      NewWARNING : Bool;   // NewWARNING
      "E-Stop BWT" : Bool;   // E-Stop BWT
      "Mask Interlocks" : Bool;   // Mask Valve Lineup Interlocks for IGG when GCU Shutting Down
      "CV403 Open" : Bool;   // Ctrl from PGC purge FB
      "CV403 Modulate Cmd" : Bool;   // Ctrl from PGC purge FB
      "CV431 Open Cmd" : Bool;   // Ctrl from PGC purge FB
      "CAB Start Cmd" : Bool;   // Ctrl from PGC purge FB
      "CAB RPM Cmd" : Real;   // Ctrl from PGC purge FB
      "CV401 Open Cmd" : Bool;   // Ctrl from PGC purge FB
   END_VAR
BEGIN
END_DATA_BLOCK

DATA_BLOCK "51_SLAVE_STATUS"   // DB51
TITLE = Slave Status Data
{ S7_Optimized_Access := 'FALSE' }
AUTHOR : JRS
VERSION : 0.1
// Data area for status from slave PLC
   VAR
      PIT112_SCALED : Real;   // IA Inlet pressure
      CV203_CNTRL : Real;   // Main fuel reg Valve Control
      PIT204_SCALED : Real;   // IGG Inlet fuel pressure
      CRNT_MODE : Int := 1;   // 1 = Auto, 2 = Man, 3 = FatAuto, 4 = FatMan
      HEART_BEAT : Bool;   // Heartbeat
      AUT_SEQ_RNG : Bool;   // Auto sequence running
      VLVS_AT_INIT : Bool;   // All valves in initial state
      P301_ENBLD : Bool;   // P301 enabled input sent from BC
      P301_TRIPPED : Bool;   // P301 tripped input sent from BC
      TS006_OK : Bool;   // TS006 Is healthy
      TS403_OK : Bool;   // TS403 Is healthy
      LS001_OK : Bool;   // LS001 Is healthy
      E131_RUNNING : Bool;   // E131 Running
      BC_SEQ_STARTED : Bool;   // BC Sequence confirmed as started
      PILOT_BURNER_ACTV : Bool;   // Pilot burn confirmed as active
      PILOT_PURGE_DN : Bool;   // Pilot burner purge completed
      RAMPING_O2_ACTV : Bool;   // Ramping of O2 is active
      O2_LVL_OK : Bool;   // O2 Level within specification
      SHTNG_DN_CNF : Bool;   // Shutting down confirmed
      O2_CNTRL_STPD : Bool;   // O2 Control modulation stopped
      BURNS_STOPPED : Bool;   // Confirmation burners are off
      CV127_CLOSED : Bool;   // CV127 Closed status
      CV203_CLOSED : Bool;   // CV203 Closed status
      CV111_CLOSED : Bool;   // CV111 Closed status
      BC_SD_DONE : Bool;   // BC Shutdown sequence done
      BC_ALARM : Bool;   // 1 = BC Alarm state, 0 = Not
      MAA_PRES_IN_RNG : Bool;   // PIT113 Main atom air pressure within range
      "FD001FDU Healthy" : Bool;   // FDU Healthy
      "FS 317 Healthy" : Bool;   // Jacket Cooling Water Flow Switch
      "PIT 204 Healthy" : Bool;   // PIT 204 Healthy
      "FS 320 Healthy" : Bool;   // FS 320 Healthy
      Warnings : Bool;   // Warnings
      "PIT 112 Healthy" : Bool;   // PIT 112 Healthy
      MAIN_BURNER_ACTV : Bool;   // MAIN_BURNER_ACTV
      "BC New ALARM" : Bool;   // New BC Alarm
      "BC New WARNING" : Bool;   // New BC Warning
      P305_ENBLD : Bool;   // P305 enabled input sent from BC
      P305_TRIPPED : Bool;   // P305 tripped input sent from BC
      P305_PRSNT : Bool;   // P305_PRSNT
      SPR_18_3 : Bool;   // Spare bit
      SPR_18_4 : Bool;   // Spare bit
      SPR_18_5 : Bool;   // Spare bit
      SPR_18_6 : Bool;   // Spare bit
      SPR_18_7 : Bool;   // Spare bit
   END_VAR
BEGIN
END_DATA_BLOCK

DATA_BLOCK "55_STATUS_DATA"   // DB55
TITLE = Status Data
{ S7_Optimized_Access := 'FALSE' }
AUTHOR : JRS
VERSION : 0.1
// Data area for status to master PLC
   VAR
      HEART_BEAT : Bool;   // Heartbeat
      AUT_SEQ_RNG : Bool;   // Auto sequence running
      CRNT_MODE : Int := 1;   // 1 = Auto, 2 = Man, 3 = FatAuto, 4 = FatMan
      STARTING : Bool;   // IGG Is starting
      O2_LVL_OK : Bool;   // O2 Level within specification
      RUNNING : Bool;   // Running
      VLVS_AT_INIT : Bool;   // 1 = Valves at initial, 0 = Not
      ESTOP_OK : Bool;   // 1 = OK, 0 = Estop active
      IGG_ALARM : Bool;   // 1 = IGG Alarm state, 0 = Not
      P305_ENBLD : Bool;   // P305 enabled input sent from BC
      P305_TRIPPED : Bool;   // P305 tripped input sent from BC
      CV401_OPN : Bool;   // CV401 Open
      CV401_CLSD : Bool;   // CV401 Closed
      P301_ENBLD : Bool;   // P305 enabled input sent from BC
      CV311_OPN : Bool;   // CV311 Open
      CV311_CLSD : Bool;   // CV311 CLosed
      CV322_OPN : Bool;   // CV322 Open
      CV322_CLSD : Bool;   // CV322 Closed
      Reset_Alarms : Bool;   // Reset_Alarms
      P305_PRSNT : Bool;
      ALARM_PRSNT : Bool;   // Alarms to master PLC
      "CV403 Less 50%" : Bool;
      "BWT Mode Selected" : Bool;
      "CB Mode Selected" : Bool;
      CV321_CLSD : Bool;
      "CAB Started" : Bool;
      "CV403 Opening" : Real;
      "CV431 Opened" : Bool;
      "IGG Stoped" : Bool;
   END_VAR
BEGIN
END_DATA_BLOCK

DATA_BLOCK "56_SLAVE_CMNDS"   // DB56
TITLE = Slave Command Data
{ S7_Optimized_Access := 'FALSE' }
AUTHOR : JRS
VERSION : 0.1
// Data area for commands to slave PLC
   VAR
      CRNT_MODE : Int := 1;   // 1 = Auto, 2 = Man, 3 = FatAuto, 4 = FatMan
      HEART_BEAT : Bool;   // Heartbeat
      ESTOP_OK : Bool;   // 1 = OK, 0 = Estop active
      RST_AUT_SEQ : Bool;   // Reset automatic sequence
      RUN_E131 : Bool;   // IA Compressor demand
      RUN_P301 : Bool;   // 1 = Run, 0 = Not
      RUN_BC_SEQ : Bool;   // 1 = Start command. 0 = Not
      PB_STS_CNFMD : Bool;   // Pilot burn status confirmed by IGG
      CRG_BLNK_MODE : Bool;   // 1 = Cargon blanketing mode, 0 = Not
      RUN_BC_O2_RAMP : Bool;   // 1 = Run ramp, 0 = Not
      BC_SD_CMND : Bool;   // 1 = Run, 0 = Shutdown
      STOP_BURNS_CMND : Bool;   // 1 = Burners off, 0 = Not
      CLS_CV127_CMND : Bool;   // 1 = Close, 0 = Not
      CLS_CV203_CMND : Bool;   // 1 = Close, 0 = Not
      CLS_CV111_CMND : Bool;   // 1 = Close, 0 = Not
      IGG_ALARM : Bool;   // 1 = IGG Alarm state, 0 = Not
      RUN_P305 : Bool;   // Fresh water pump demand
      CV403_OPEN : Bool;   // 1 = Valve is open, 0 = Not
      "E 500A RUN" : Bool;   // Fuel Pump 1 Enabled
      "E 500B RUN" : Bool;   // Fuel Pump 2 Enabled
      "TIT 360 Healthy" : Bool;   // Outlet CSW Temp TIT360
      "TIT 401 Healthy" : Bool;   // IG Temp
      "PIT 316 Healthy" : Bool;   // Outlet CSW Pressure
      RST_LOCKOUT : Bool;   // Reset of alarms
      "CA Blower Running" : Bool;   // E139-MCCP/6TA1
      Alarm_Reset : Bool;   // Alarm_Reset
      BWT_MODE : Bool;
      "P301 PRSNT" : Bool;
      "TIT 315 Healthy" : Bool;   // PIT 315 Healthy
      SFTY_SYS_IL : Bool;   // SFTY_SYS_IL
      "Master Stop" : Bool;   // Master Stop
      "CV401 Closed" : Bool;   // CV401 Closed
      SPR_5_7 : Bool;   // Spare bool
      IGG_CRNT_STEP : Int;   // IGG Current Step
   END_VAR
BEGIN
END_DATA_BLOCK

DATA_BLOCK "58_COMMS_DATE_TIME"   // DB58
{ S7_Optimized_Access := 'FALSE' }
VERSION : 0.1
   VAR
      SYSTEM_TIME : DTL;
      LOCAL_TIME : DTL;
   END_VAR
BEGIN
END_DATA_BLOCK

DATA_BLOCK "59_COMMS_HEALTH_DATA"   // DB59
TITLE = Communications Health Data
{ S7_Optimized_Access := 'TRUE' }
AUTHOR : JRS
VERSION : 0.1
// Data area for communications health determination
   VAR
      CLOCK_POS_EDGE : Bool;   // Edge bit
      CLOCK_NEG_EDGE : Bool;   // Edge bit
      MSTR_TRUE_TMR : TON_TIME;
      MSTR_FALSE_TMR : TON_TIME;
      SLAVE_TRUE_TMR : TON_TIME;
      SLAVE_FALSE_TMR : TON_TIME;
      MSTR_HB_MISSING : Bool;   // Heatbeat missing flag
      SLAVE_HB_MISSING : Bool;   // Heartbeat missing flag
      "IGG HMI HB" : Bool;
      "IGG HMI HB MISSING" : Bool;
      "IGG HMI HB ON TIMER" : TON_TIME;
      "IGG HMI HB OFF TIMER" : TON_TIME;
      "CCR HMI HB" : Bool;
      "CCR HMI HB MISSING" : Bool;
      "CCR HMI HB ON TIMER" : TON_TIME;
      "CCR HMI HB OFF TIMER" : TON_TIME;
      "BRIGE HMI HB" : Bool;
      "BRIGE HMI HB MISSING" : Bool;
      "BRIGE HMI HB ON TIMER" : TON_TIME;
      "BRIGE HMI HB OFF TIMER" : TON_TIME;
      "GET HEALTH" : Bool;
      "PUT HEALTH" : Bool;
   END_VAR
BEGIN
   MSTR_FALSE_TMR.PT := T#2s;
   MSTR_TRUE_TMR.PT := T#2s;
   SLAVE_TRUE_TMR.PT := T#2s;
   SLAVE_FALSE_TMR.PT := T#2s;
END_DATA_BLOCK

// folder: 60 - 69 Alarm & Status Handling

DATA_BLOCK "503_ALARM CHCK_DB_1"   // DB2
{ S7_Optimized_Access := 'TRUE' }
VERSION : 0.1
// stored: InstanceOfName 503_ALARM CHCK
"503_ALARM CHCK"
BEGIN
END_DATA_BLOCK

DATA_BLOCK "60_Alarm_Data"   // DB60
{ S7_Optimized_Access := 'FALSE' }
VERSION : 0.1
   VAR
      IGG_ALARM_WORD_01 : Word;
      IGG_ALARM_WORD_02 : Word;
      IGG_ALARM_WORD_03 : Word;
      IGG_ALARM_WORD_04 : Word;
      IGG_ALARM_WORD_05 : Word;
      IGG_ALARM_WORD_06 : Word;
      IGG_ALARM_WORD_07 : Word;
      IGG_ALARM_WORD_08 : Word;
      IGG_ALARM_WORD_09 : Word;
      IGG_ALARM_WORD_10 : Word;
      IGG_ALARM_WORD_11 : Word;
      IGG_ALARM_WORD_12 : Word;
      IGG_ALARM_WORD_13 : Word;
      IGG_ALARM_WORD_14 : Word;
      IGG_ALARM_WORD_15 : Word;
      IGG_ALARM_WORD_16 : Word;
      ALRM_PRSNT : Bool;
   END_VAR
BEGIN
END_DATA_BLOCK
